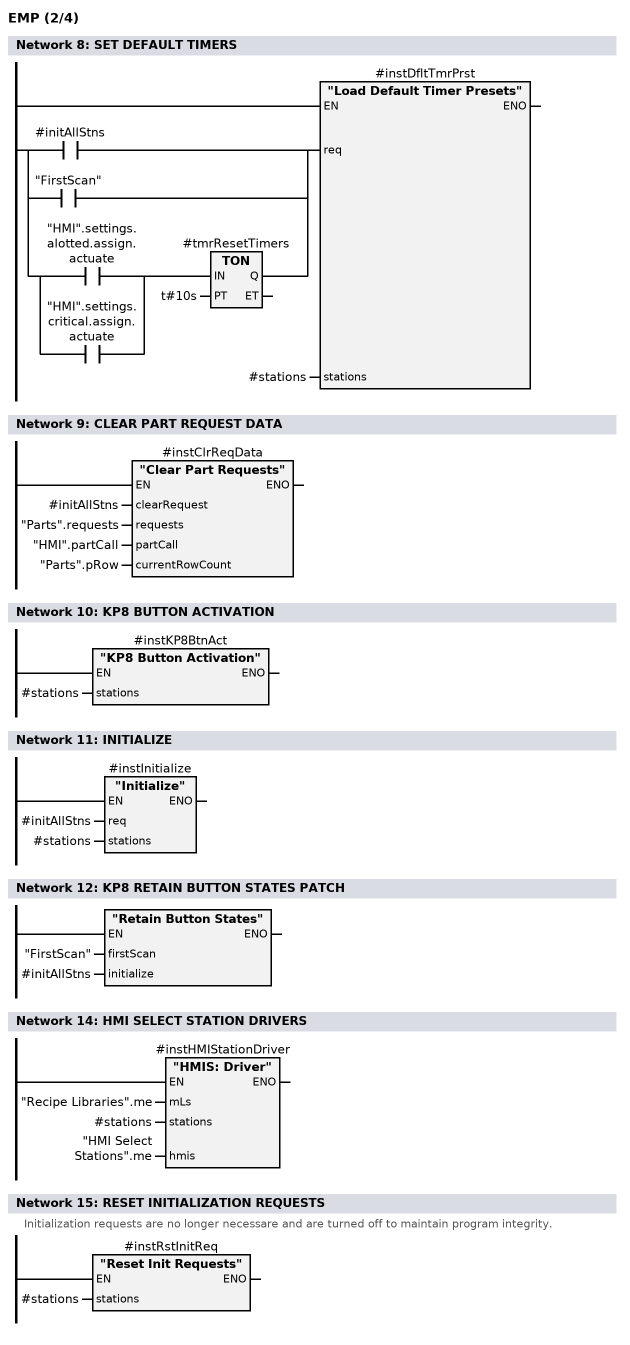
   #tmrResetTimers(IN := "HMI".settings.alotted.assign.actuate OR "HMI".settings.critical.assign.actuate,   // TON
                   PT := t#10s);
   #instDfltTmrPrst(req := #initAllStns OR "FirstScan" OR #tmrResetTimers.Q, stations := #stations);   // "Load Default Timer Presets"
END_REGION

REGION Network 9: CLEAR PART REQUEST DATA
   RUNG wire#powerrail
      #instClrReqData(clearRequest := #initAllStns, requests := "Parts".requests, partCall := "HMI".partCall, currentRowCount := "Parts".pRow)
   END_RUNG
   // the same network as SCL:
   #instClrReqData(clearRequest := #initAllStns,   // "Clear Part Requests"
                   requests := "Parts".requests,
                   partCall := "HMI".partCall,
                   currentRowCount := "Parts".pRow);
END_REGION

REGION Network 10: KP8 BUTTON ACTIVATION
   RUNG wire#powerrail
      #instKP8BtnAct(stations := #stations)
   END_RUNG
   // the same network as SCL:
   #instKP8BtnAct(stations := #stations);   // "KP8 Button Activation"
END_REGION

REGION Network 11: INITIALIZE
   RUNG wire#powerrail
      #instInitialize(req := #initAllStns, stations := #stations)
   END_RUNG
   // the same network as SCL:
   #instInitialize(req := #initAllStns, stations := #stations);   // "Initialize"
END_REGION

REGION Network 12: KP8 RETAIN BUTTON STATES PATCH
   RUNG wire#powerrail
      "Retain Button States"(firstScan := "FirstScan", initialize := #initAllStns)
   END_RUNG
   // the same network as SCL:
   "Retain Button States"(firstScan := "FirstScan", initialize := #initAllStns);
END_REGION

REGION Network 13 (SCL): KP8 DRIVER CALLS
   REGION "LOOP THROUGH STATIONS"
       FOR #i := 0 TO "stnCount" DO
           CASE #i OF
               0..24, 30:
                   #instKP8Drvs[#i](btnIn := #stations.me[#i].kp8In,
                                    hardInit := #stations.me[#i].init.hard,
                                    softInit := #stations.me[#i].init.soft,
                                    btn0Activate := #stations.me[#i].kp8Config.activate[0],
                                    btn0Mode := #stations.me[#i].kp8Config.mode[0],
                                    btn0Group := #stations.me[#i].kp8Config.group[0],
                                    btn0Flash := #stations.me[#i].kp8Config.flash[0],
                                    btn0ColorOn1 := #stations.me[#i].kp8Config.colorOn1[0],
                                    btn0ColorOn2 := #stations.me[#i].kp8Config.colorOn2[0],
                                    btn0ColorOff := #stations.me[#i].kp8Config.colorOff[0],
                                    btn1Activate := #stations.me[#i].kp8Config.activate[1],
                                    btn1Mode := #stations.me[#i].kp8Config.mode[1],
                                    btn1Group := #stations.me[#i].kp8Config.group[1],
                                    btn1Flash := #stations.me[#i].kp8Config.flash[1],
                                    btn1ColorOn1 := #stations.me[#i].kp8Config.colorOn1[1],
                                    btn1ColorOn2 := #stations.me[#i].kp8Config.colorOn2[1],
                                    btn1ColorOff := #stations.me[#i].kp8Config.colorOff[1],
                                    btn2Activate := #stations.me[#i].kp8Config.activate[2],
                                    btn2Mode := #stations.me[#i].kp8Config.mode[2],
                                    btn2Group := #stations.me[#i].kp8Config.group[2],
                                    btn2Flash := #stations.me[#i].kp8Config.flash[2],
                                    btn2ColorOn1 := #stations.me[#i].kp8Config.colorOn1[2],
                                    btn2ColorOn2 := #stations.me[#i].kp8Config.colorOn2[2],
                                    btn2ColorOff := #stations.me[#i].kp8Config.colorOff[2],
                                    btn3Activate := #stations.me[#i].kp8Config.activate[3],
                                    btn3Mode := #stations.me[#i].kp8Config.mode[3],
                                    btn3Group := #stations.me[#i].kp8Config.group[3],
                                    btn3Flash := #stations.me[#i].kp8Config.flash[3],
                                    btn3ColorOn1 := #stations.me[#i].kp8Config.colorOn1[3],
                                    btn3ColorOn2 := #stations.me[#i].kp8Config.colorOn2[3],
                                    btn3ColorOff := #stations.me[#i].kp8Config.colorOff[3],
                                    btn4Activate := #stations.me[#i].kp8Config.activate[4],
                                    btn4Mode := #stations.me[#i].kp8Config.mode[4],
                                    btn4Group := #stations.me[#i].kp8Config.group[4],
                                    btn4Flash := #stations.me[#i].kp8Config.flash[4],
                                    btn4ColorOn1 := #stations.me[#i].kp8Config.colorOn1[4],
                                    btn4ColorOn2 := #stations.me[#i].kp8Config.colorOn2[4],
                                    btn4ColorOff := #stations.me[#i].kp8Config.colorOff[4],
                                    btn5Activate := #stations.me[#i].kp8Config.activate[5],
                                    btn5Mode := #stations.me[#i].kp8Config.mode[5],
                                    btn5Group := #stations.me[#i].kp8Config.group[5],
                                    btn5Flash := #stations.me[#i].kp8Config.flash[5],
                                    btn5ColorOn1 := #stations.me[#i].kp8Config.colorOn1[5],
                                    btn5ColorOn2 := #stations.me[#i].kp8Config.colorOn2[5],
                                    btn5ColorOff := #stations.me[#i].kp8Config.colorOff[5],
                                    btn6Activate := #stations.me[#i].kp8Config.activate[6],
                                    btn6Mode := #stations.me[#i].kp8Config.mode[6],
                                    btn6Group := #stations.me[#i].kp8Config.group[6],
                                    btn6Flash := #stations.me[#i].kp8Config.flash[6],
                                    btn6ColorOn1 := #stations.me[#i].kp8Config.colorOn1[6],
                                    btn6ColorOn2 := #stations.me[#i].kp8Config.colorOn2[6],
                                    btn6ColorOff := #stations.me[#i].kp8Config.colorOff[6],
                                    btn7Activate := #stations.me[#i].kp8Config.activate[7],
                                    btn7Mode := #stations.me[#i].kp8Config.mode[7],
                                    btn7Group := #stations.me[#i].kp8Config.group[7],
                                    btn7Flash := #stations.me[#i].kp8Config.flash[7],
                                    btn7ColorOn1 := #stations.me[#i].kp8Config.colorOn1[7],
                                    btn7ColorOn2 := #stations.me[#i].kp8Config.colorOn2[7],
                                    btn7ColorOff := #stations.me[#i].kp8Config.colorOff[7],
                                    btnStatesOut => #stations.me[#i].btnStates,
                                    btnColorsOut => #stations.me[#i].kp8Out);
               ELSE 
                   ;
           END_CASE;

       END_FOR;
   END_REGION
END_REGION

REGION Network 14: HMI SELECT STATION DRIVERS
   RUNG wire#powerrail
      #instHMIStationDriver(mLs := "Recipe Libraries".me, stations := #stations, hmis := "HMI Select Stations".me)
   END_RUNG
   // the same network as SCL:
   #instHMIStationDriver(mLs := "Recipe Libraries".me, stations := #stations, hmis := "HMI Select Stations".me);   // "HMIS: Driver"
END_REGION

REGION Network 15: RESET INITIALIZATION REQUESTS
   // Initialization requests are no longer necessare and are turned off to maintain program integrity.
   RUNG wire#powerrail
      #instRstInitReq(stations := #stations)
   END_RUNG
   // the same network as SCL:
   #instRstInitReq(stations := #stations);   // "Reset Init Requests"
END_REGION

REGION Network 16: BARCODE SCREEN
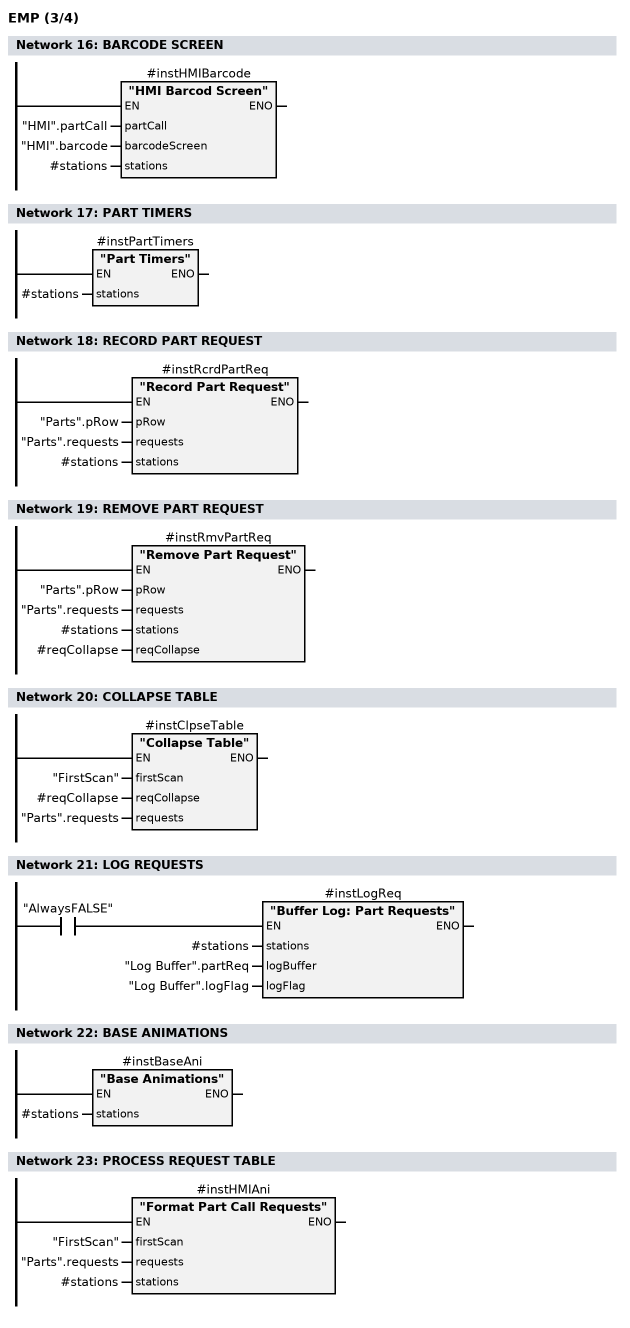
   RUNG wire#powerrail
      #instHMIBarcode(partCall := "HMI".partCall, barcodeScreen := "HMI".barcode, stations := #stations)
   END_RUNG
   // the same network as SCL:
   #instHMIBarcode(partCall := "HMI".partCall, barcodeScreen := "HMI".barcode, stations := #stations);   // "HMI Barcod Screen"
END_REGION

REGION Network 17: PART TIMERS
   RUNG wire#powerrail
      #instPartTimers(stations := #stations)
   END_RUNG
   // the same network as SCL:
   #instPartTimers(stations := #stations);   // "Part Timers"
END_REGION

REGION Network 18: RECORD PART REQUEST
   RUNG wire#powerrail
      #instRcrdPartReq(pRow := "Parts".pRow, requests := "Parts".requests, stations := #stations)
   END_RUNG
   // the same network as SCL:
   #instRcrdPartReq(pRow := "Parts".pRow, requests := "Parts".requests, stations := #stations);   // "Record Part Request"
END_REGION

REGION Network 19: REMOVE PART REQUEST
   RUNG wire#powerrail
      #instRmvPartReq(pRow := "Parts".pRow, requests := "Parts".requests, stations := #stations, reqCollapse := #reqCollapse)
   END_RUNG
   // the same network as SCL:
   #instRmvPartReq(pRow := "Parts".pRow,   // "Remove Part Request"
                   requests := "Parts".requests,
                   stations := #stations,
                   reqCollapse := #reqCollapse);
END_REGION

REGION Network 20: COLLAPSE TABLE
   RUNG wire#powerrail
      #instClpseTable(firstScan := "FirstScan", reqCollapse := #reqCollapse, requests := "Parts".requests)
   END_RUNG
   // the same network as SCL:
   #instClpseTable(firstScan := "FirstScan", reqCollapse := #reqCollapse, requests := "Parts".requests);   // "Collapse Table"
END_REGION

REGION Network 21: LOG REQUESTS
   RUNG wire#powerrail
      Contact( "AlwaysFALSE" )
      #instLogReq(stations := #stations, logBuffer := "Log Buffer".partReq, logFlag := "Log Buffer".logFlag)
   END_RUNG
   // the same network as SCL:
   IF "AlwaysFALSE" THEN
       #instLogReq(stations := #stations, logBuffer := "Log Buffer".partReq, logFlag := "Log Buffer".logFlag);   // "Buffer Log: Part Requests"
   END_IF;
END_REGION

REGION Network 22: BASE ANIMATIONS
   RUNG wire#powerrail
      #instBaseAni(stations := #stations)
   END_RUNG
   // the same network as SCL:
   #instBaseAni(stations := #stations);   // "Base Animations"
END_REGION

REGION Network 23: PROCESS REQUEST TABLE
   RUNG wire#powerrail
      #instHMIAni(firstScan := "FirstScan", requests := "Parts".requests, stations := #stations)
   END_RUNG
   // the same network as SCL:
   #instHMIAni(firstScan := "FirstScan", requests := "Parts".requests, stations := #stations);   // "Format Part Call Requests"
END_REGION

REGION Network 24: HMI POPULATE TABLE
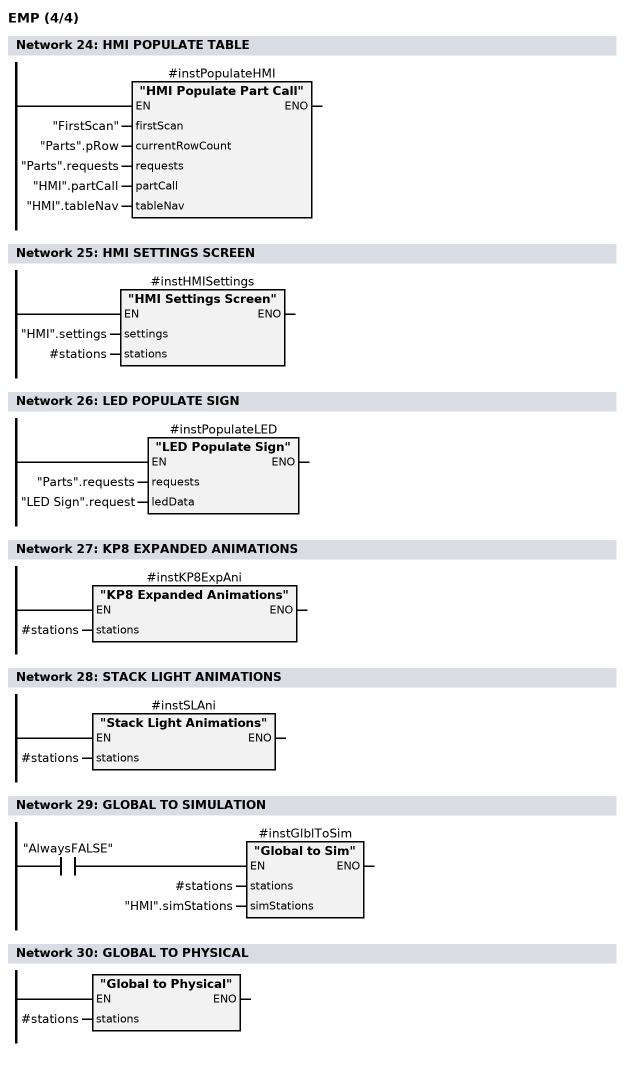
   RUNG wire#powerrail
      #instPopulateHMI(firstScan := "FirstScan", currentRowCount := "Parts".pRow, requests := "Parts".requests, partCall := "HMI".partCall, tableNav := "HMI".tableNav)
   END_RUNG
   // the same network as SCL:
   #instPopulateHMI(firstScan := "FirstScan",   // "HMI Populate Part Call"
                    currentRowCount := "Parts".pRow,
                    requests := "Parts".requests,
                    partCall := "HMI".partCall,
                    tableNav := "HMI".tableNav);
END_REGION

REGION Network 25: HMI SETTINGS SCREEN
   RUNG wire#powerrail
      #instHMISettings(settings := "HMI".settings, stations := #stations)
   END_RUNG
   // the same network as SCL:
   #instHMISettings(settings := "HMI".settings, stations := #stations);   // "HMI Settings Screen"
END_REGION

REGION Network 26: LED POPULATE SIGN
   RUNG wire#powerrail
      #instPopulateLED(requests := "Parts".requests, ledData := "LED Sign".request)
   END_RUNG
   // the same network as SCL:
   #instPopulateLED(requests := "Parts".requests, ledData := "LED Sign".request);   // "LED Populate Sign"
END_REGION

REGION Network 27: KP8 EXPANDED ANIMATIONS
   RUNG wire#powerrail
      #instKP8ExpAni(stations := #stations)
   END_RUNG
   // the same network as SCL:
   #instKP8ExpAni(stations := #stations);   // "KP8 Expanded Animations"
END_REGION

REGION Network 28: STACK LIGHT ANIMATIONS
   RUNG wire#powerrail
      #instSLAni(stations := #stations)
   END_RUNG
   // the same network as SCL:
   #instSLAni(stations := #stations);   // "Stack Light Animations"
END_REGION

REGION Network 29: GLOBAL TO SIMULATION
   RUNG wire#powerrail
      Contact( "AlwaysFALSE" )
      #instGlblToSim(stations := #stations, simStations := "HMI".simStations)
   END_RUNG
   // the same network as SCL:
   IF "AlwaysFALSE" THEN
       #instGlblToSim(stations := #stations, simStations := "HMI".simStations);   // "Global to Sim"
   END_IF;
END_REGION

REGION Network 30: GLOBAL TO PHYSICAL
   RUNG wire#powerrail
      "Global to Physical"(stations := #stations)
   END_RUNG
   // the same network as SCL:
   "Global to Physical"(stations := #stations);
END_REGION
END_FUNCTION_BLOCK

FUNCTION "Retain Button States" : Void   // FC36, SCL
{ S7_Optimized_Access := 'TRUE' }
VERSION : 0.1
   VAR_INPUT
      firstScan : Bool;
      initialize : Bool;
   END_VAR
   VAR_TEMP
      i : Int;
      j : Int;
   END_VAR
BEGIN
   FOR #i := 0 TO "stnCount" DO
           FOR #j := 0 TO "ptsPerStn" DO
               IF #firstScan THEN
                   "EMP IDB".instKP8Drvs[#i].btnStateArrayInt[#j] :=
                   "EMP IDB".stations.me[#i].btnStates[#j];
               END_IF;
               IF #initialize THEN
                   "EMP IDB".instKP8Drvs[#i].btnStateArrayInt[#j] := FALSE;
                   "EMP IDB".stations.me[#i].btnStates[#j] := FALSE;
               END_IF;
           END_FOR;
   END_FOR;
END_FUNCTION

ORGANIZATION_BLOCK "Main"   // OB1, LAD, ProgramCycle
TITLE = "Main Program Sweep (Cycle)"
{ S7_Optimized_Access := 'TRUE' }
VERSION : 0.1
   VAR_INPUT
      Initial_Call : Bool;   // Initial call of this OB
      Remanence : Bool;   // =True, if remanent data are available
   END_VAR
BEGIN

REGION Network 1
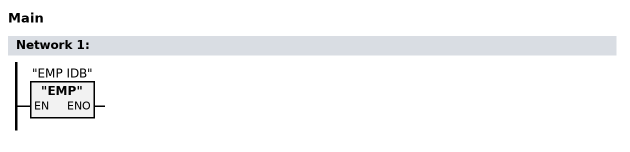
   RUNG wire#powerrail
      "EMP IDB"()
   END_RUNG
   // the same network as SCL:
   "EMP IDB"();   // "EMP"
END_REGION
END_ORGANIZATION_BLOCK

// folder: Global/Physical

FUNCTION "Physical to Global" : Void   // FC1, LAD
{ S7_Optimized_Access := 'TRUE' }
VERSION : 0.1
   VAR_IN_OUT
      stations : "Stations";
   END_VAR
   VAR_TEMP
      i : Int;
      kp8In : DWord;
   END_VAR
BEGIN

REGION Network 1 (SCL): MAIN LOOP
   FOR #i := 0 TO "stnCount" DO

       CASE #i OF
           "VOLVO 16 01":
               #kp8In := "VOLVO 16 01 KP8 In";
           "VOLVO 16 02":
               #kp8In := "VOLVO 16 02 KP8 In";
           "VOLVO 16 03":
               #kp8In := "VOLVO 16 03 KP8 In";
           "VOLVO 16 04":
               #kp8In := "VOLVO 16 04 KP8 In";
           "VOLVO 16 05":
               #kp8In := "VOLVO 16 05 KP8 In";
           "VOLVO 16 06":
               #kp8In := "VOLVO 16 06 KP8 In";
           "VOLVO 16 07":
               #kp8In := "VOLVO 16 07 KP8 In";
           "VOLVO 16 08":
               #kp8In := "VOLVO 16 08 KP8 In";
           "VOLVO 16 09":
               #kp8In := "VOLVO 16 09 KP8 In";
           "VOLVO 16 10":
               #kp8In := "VOLVO 16 10 KP8 In";
           "VOLVO 16 11":
               #kp8In := "VOLVO 16 11 KP8 In";
           "CHM 01":
               #kp8In := "CHM 01 KP8 In";
           "CHM 02":
               #kp8In := "CHM 02 KP8 In";
           "CHM 03":
               #kp8In := "CHM 03 KP8 In";
           "CHM 04":
               #kp8In := "CHM 04 KP8 In";
           "CHM 05":
               #kp8In := "CHM 05 KP8 In";
           "CDO 01":
               #kp8In := "CDO 01 KP8 In";
           "CDO 02":
               #kp8In := "CDO 02 KP8 In";
           "CDO 03":
               #kp8In := "CDO 03 KP8 In";
           "BFL 01":
               #kp8In := "BFL 01 KP8 In";
           "BFL 02":
               #kp8In := "BFL 02 KP8 In";
           "BFL 03":
               #kp8In := "BFL 03 KP8 In";
           "LGS 01":
               #kp8In := "LGS 01 KP8 In";
           "LGS 02":
               #kp8In := "LGS 02 KP8 In";
           "LGS 03":
               #kp8In := "LGS 03 KP8 In";
           "CV 01":
               #kp8In := "CV 01 KP8 In";
           "CV 02":
               #kp8In := "CV 02 KP8 In";
           "CV 03":
               #kp8In := "CV 03 KP8 In";
           "CV 04":
               #kp8In := "CV 04 KP8 In";
           "PC 01":
               #kp8In := "PC 01 KP8 In"; 
           "PC 02":
               #kp8In := "PC 02 KP8 In";
       END_CASE;

       #stations.me[#i].kp8In := #kp8In.%B3;

   END_FOR;
END_REGION
END_FUNCTION

FUNCTION "Global to Physical" : Void   // FC5, LAD
{ S7_Optimized_Access := 'TRUE' }
VERSION : 0.1
   VAR_IN_OUT
      stations : "Stations";
   END_VAR
   VAR_TEMP
      i : Int;
      j : Int;
      IO : DWord;
      "KP8 In" : DWord;
      "KP8 Out" : DWord;
      Card : Int;
      stnCount : Int;
   END_VAR
BEGIN

REGION Network 1 (SCL): MAIN LOOP
   FOR #i := 0 TO "stnCount" DO

       #IO := #stations.me[#i].stackLightOut;
       #"KP8 Out" := #stations.me[#i].kp8Out;

       CASE #i OF
           "VOLVO 16 01":
               "VOLVO 16 01 IO" := #IO;
               "VOLVO 16 01 KP8 Out" := #"KP8 Out";
           "VOLVO 16 02":
               "VOLVO 16 02 IO" := #IO;
               "VOLVO 16 02 KP8 Out" := #"KP8 Out";
           "VOLVO 16 03":
               "VOLVO 16 03 IO" := #IO;
               "VOLVO 16 03 KP8 Out" := #"KP8 Out";
           "VOLVO 16 04":
               "VOLVO 16 04 IO" := #IO;
               "VOLVO 16 04 KP8 Out" := #"KP8 Out";
           "VOLVO 16 05":
               "VOLVO 16 05 IO" := #IO;
               "VOLVO 16 05 KP8 Out" := #"KP8 Out";
           "VOLVO 16 06":
               "VOLVO 16 06 IO" := #IO;
               "VOLVO 16 06 KP8 Out" := #"KP8 Out";
           "VOLVO 16 07":
               "VOLVO 16 07 IO" := #IO;
               "VOLVO 16 07 KP8 Out" := #"KP8 Out";
           "VOLVO 16 08":
               "VOLVO 16 08 IO" := #IO;
               "VOLVO 16 08 KP8 Out" := #"KP8 Out";
           "VOLVO 16 09":
               "VOLVO 16 09 IO" := #IO;
               "VOLVO 16 09 KP8 Out" := #"KP8 Out";
           "VOLVO 16 10":
               "VOLVO 16 10 IO" := #IO;
               "VOLVO 16 10 KP8 Out" := #"KP8 Out";
           "VOLVO 16 11":
               "VOLVO 16 11 IO" := #IO;
               "VOLVO 16 11 KP8 Out" := #"KP8 Out";
           "CHM 01":
               "CHM 01 IO" := #IO;
               "CHM 01 KP8 Out" := #"KP8 Out";
           "CHM 02":
               "CHM 02 IO" := #IO;
               "CHM 02 KP8 Out" := #"KP8 Out";
           "CHM 03":
               "CHM 03 IO" := #IO;
               "CHM 03 KP8 Out" := #"KP8 Out";
           "CHM 04":
               "CHM 04 IO" := #IO;
               "CHM 04 KP8 Out" := #"KP8 Out";
           "CHM 05":
               "CHM 05 IO" := #IO;
               "CHM 05 KP8 Out" := #"KP8 Out";
           "CDO 01":
               "CDO 01 IO" := #IO;
               "CDO 01 KP8 Out" := #"KP8 Out";
           "CDO 02":
               "CDO 02 IO" := #IO;
               "CDO 02 KP8 Out" := #"KP8 Out";
           "CDO 03":
               "CDO 03 IO" := #IO;
               "CDO 03 KP8 Out" := #"KP8 Out";
           "BFL 01":
               "BFL 01 IO" := #IO;
               "BFL 01 KP8 Out" := #"KP8 Out";
           "BFL 02":
               "BFL 02 IO" := #IO;
               "BFL 02 KP8 Out" := #"KP8 Out";
           "BFL 03":
               "BFL 03 IO" := #IO;
               "BFL 03 KP8 Out" := #"KP8 Out";
           "LGS 01":
               "LGS 01 IO" := #IO;
               "LGS 01 KP8 Out" := #"KP8 Out";
           "LGS 02":
               "LGS 02 IO" := #IO;
               "LGS 02 KP8 Out" := #"KP8 Out";
           "LGS 03":
               "LGS 03 IO" := #IO;
               "LGS 03 KP8 Out" := #"KP8 Out";
           "CV 01":
               "CV 01 IO" := #IO;
               "CV 01 KP8 Out" := #"KP8 Out";
           "CV 02":
               "CV 02 IO" := #IO;
               "CV 02 KP8 Out" := #"KP8 Out";
           "CV 03":
               "CV 03 IO" := #IO;
               "CV 03 KP8 Out" := #"KP8 Out";
           "CV 04":
               "CV 04 IO" := #IO;
               "CV 04 KP8 Out" := #"KP8 Out";
           "PC 01":
               "PC 01 IO" := #IO;
               "PC 01 KP8 Out" := #"KP8 Out";
           "PC 02":
               "PC 02 IO" := #IO;
               "PC 02 KP8 Out" := #"KP8 Out";

       END_CASE;

   END_FOR;
END_REGION
END_FUNCTION

// folder: HMI Stations

FUNCTION_BLOCK "HMIS: Driver"   // FB32, LAD
{ S7_Optimized_Access := 'TRUE' }
VERSION : 0.1
   VAR_INPUT
      mLs : "Recipe: Libraries";
   END_VAR
   VAR_IN_OUT
      stations : "Stations";
      hmis : Array[0.."hmiStnCount"] of "HSS: Compressed";
   END_VAR
   VAR
      recipeSelector : Array[0.."hmiStnCount"] of Int;
      r1 : Array[0.."hmiStnCount"] of DInt;
      instsHSSMenuSelect : Array[0.."hmiStnCount"] of "HMIS: Recipe Selection";
      instsHSSPartSelect : Array[0.."hmiStnCount"] of "HMIS: Part Selection";
   END_VAR
   VAR_TEMP
      i : Int;
   END_VAR
   VAR CONSTANT
      hssOffset : Int := 25;
   END_VAR
BEGIN

REGION Network 1 (SCL): TEMPLATE SCREENS
   FOR #i := 0 TO "hmiStnCount" DO
       "HMIS: Template"(menuLibrary := #mLs.stations[#i + #hssOffset],
                       menuSelector := #recipeSelector[#i],
                       tmplt := #hmis[#i].scrnTmplt);
       #instsHSSMenuSelect[#i](lib := #mLs.stations[#i + #hssOffset],
                               slctScreen := #hmis[#i].scrnSlctMn,
                               r1 := #r1[#i],
                               station := #stations.me[#i + #hssOffset],
                               recipeSelector := #recipeSelector[#i]);
       #instsHSSPartSelect[#i](recipeNum:= #recipeSelector[#i],
                              lib:=#mLs.stations[#i + #hssOffset],
                              slctScreen:=#hmis[#i].scrnSlctPrt,
                              station:=#stations.me[#i + #hssOffset]);

   END_FOR;
END_REGION
END_FUNCTION_BLOCK

FUNCTION_BLOCK "HMIS: Part Selection"   // FB33, SCL
{ S7_Optimized_Access := 'TRUE' }
VERSION : 0.1
   VAR_INPUT
      recipeNum : Int;
      lib : "Recipe: Library";
   END_VAR
   VAR_IN_OUT
      slctScreen : "HSS: Part Selection Screen";
      station : "Station";
   END_VAR
   VAR
      oldBtnsIn : Array[0..31] of Bool;
   END_VAR
   VAR_TEMP
      eval : "HSS: Part Selection Screen";
      i : Int;
      btnsIn : Array[0..31] of Bool;
      btnStates : Array[0.."ptsPerStn"] of Bool;
   END_VAR
BEGIN
   #eval := #slctScreen;


   SCATTER(IN := #slctScreen.pbs ,
           OUT => #btnsIn);
   #btnStates := #station.btnStates;


   FOR #i := 0 TO "ptsPerStn" DO
       IF #btnsIn[#i] AND #btnsIn[#i] <> #oldBtnsIn[#i] THEN
           #btnStates[#i] := NOT #btnStates[#i];
       END_IF;
   END_FOR;


   FOR #i := 0 TO "ptsPerStn" DO
       "Part Select Button"(recipeNum := #recipeNum,
                            lib := #lib,
                            actuate := #btnsIn[#i],
                            btnNum := #i,
                            stn:= #station,
                            partSelectScreen := #eval);
   END_FOR;


   #station.btnStates := #btnStates;
   #oldBtnsIn := #btnsIn;
   #slctScreen := #eval;
END_FUNCTION_BLOCK

FUNCTION_BLOCK "HMIS: Recipe Selection"   // FB35, SCL
{ S7_Optimized_Access := 'TRUE' }
VERSION : 0.1
   VAR_INPUT
      lib : "Recipe: Library";
   END_VAR
   VAR_IN_OUT
      slctScreen : "HSS: Menu Selection Screen";
      r1 : DInt;
      recipeSelector : Int;
      station : "Station";
   END_VAR
   VAR
      old : Struct
         navPress : Bool;
      END_STRUCT;
      instTableNavigation : "Table Navigatio";
   END_VAR
   VAR_TEMP
      eval : "HSS: Menu Selection Screen";
      pbs : Array[0..#pbFlagCnt] of Bool;
      POS : DInt;
      status : DInt;
      i : Int;
      btnNum : Int;
      pRowVisLbl : Int;
      pRowInvisLbl : Int;
      pRecipeInvisLbl : Int;
      pRecipeVisLbl : Int;
      pRecipeLib : Int;
      pRowTxt : Int;
      pRecipeTxt : Int;
      shifter : DWord;
      btnsAsBool : Array[0..31] of Bool;
      rows : Array[0..99] of DInt;
      offset : DInt;
      navPress : Bool;
      selPress : Bool;
      maxRows : DInt;
      tmrReal : Real;
      partNumber : WString;
   END_VAR
   VAR CONSTANT
      pbFlagCnt : Int := 31;
      btnCnt : Int := 5;
      navMask : DWord := 16#0000_003F;
      visRows : DInt := 6;
      home : DInt := -1000;
      end : DInt := -2000;
      alotted : Real := 1800.0;
      critical : Real := 300.0;
   END_VAR
BEGIN
   REGION "INITITALIZE LOCALS"

       #eval := #slctScreen;
       #maxRows := #lib.size;
       SCATTER(IN := #eval.pbs,
               OUT => #btnsAsBool);

   END_REGION


   REGION "GET RECIPE SELECTION PRESS" 

       REGION "GET RECIPE SELECTOR NUMBER"

           FOR #i := 6 TO 31 DO
               IF #btnsAsBool[#i] THEN

                   #recipeSelector := DINT_TO_INT(#r1) + #i - 6;

                   IF #recipeSelector > #maxRows -1 THEN
                       #recipeSelector := #recipeSelector - DINT_TO_INT(#maxRows);
                   END_IF;

                   IF #recipeSelector < 0 THEN
                       #recipeSelector := DINT_TO_INT(#maxRows) + #recipeSelector;
                   END_IF;

                   #selPress := TRUE;
                   EXIT;
               END_IF;
           END_FOR;

       END_REGION


       FOR #i := 0 TO "ptsPerStn" DO
           #station.partNumbers[#i] := #lib.raw[#recipeSelector, #i];
           IF #i = 1 THEN
               #station.partNumbers[#i] := WSTRING#'DUNNAGE';
           END_IF;

       END_FOR;

       REGION "SET DEFAULT TIMERS"
           FOR #i := 0 TO "ptsPerStn" DO

               REGION "COPY TO LOCAL"
                   #partNumber := #station.partNumbers[#i];
               END_REGION

               REGION "IF BUTTON HAS ASSOCIATED PN"
                   IF LEN(#partNumber) <> 0 THEN

                       REGION "COPY TO LOCAL"
                           #tmrReal := #station.presetTime.allotted[#i];
                       END_REGION

                       REGION "ON NO TIME ENTERED"
                           IF #tmrReal = 0.0 THEN

                               REGION "ASSIGN ALLOTTED VALUES"
                                   #station.presetTime.allotted[#i] := #alotted;
                               END_REGION

                           END_IF;
                       END_REGION

                       REGION "COPY TO LOCAL"
                           #tmrReal := #station.presetTime.critical[#i];
                       END_REGION

                       REGION "ON NO TIME ENTERED"
                           IF #tmrReal = 0.0 THEN

                               REGION "ASSIGN CRITICAL VALUES"
                                   #station.presetTime.critical[#i] := #critical;
                               END_REGION

                           END_IF;
                       END_REGION

                   END_IF;
               END_REGION

               REGION "IF BUTTON HAS NO ASSOCIATED PN"
                   IF LEN(#partNumber) = 0 THEN

                       REGION "COPY TO LOCAL"
                           #tmrReal := #station.presetTime.allotted[#i];
                       END_REGION

                       REGION "ON NO TIME ENTERED"
                           IF #tmrReal <> 0.0 THEN

                               REGION "ASSIGN ALLOTTED VALUES"
                                   #station.presetTime.allotted[#i] := 0.0;
                               END_REGION

                           END_IF;
                       END_REGION

                       REGION "COPY TO LOCAL"
                           #tmrReal := #station.presetTime.critical[#i];
                       END_REGION

                       REGION "ON NO TIME ENTERED"
                           IF #tmrReal <> 0.0 THEN

                               REGION "ASSIGN CRITICAL VALUES"
                                   #station.presetTime.critical[#i] := 0.0;
                               END_REGION

                           END_IF;
                       END_REGION

                   END_IF;
               END_REGION


           END_FOR;
       END_REGION

   END_REGION


   REGION "TABLE NAVIGATION"
       IF #maxRows > #visRows THEN
           IF #eval.pbs.%X0 THEN
               #offset := #home;
           END_IF;
           IF #eval.pbs.%X1 THEN
               #offset := -1 * #visRows;
           END_IF;
           IF #eval.pbs.%X2 THEN
               #offset := -1;
           END_IF;
           IF #eval.pbs.%X3 THEN
               #offset := 1;
           END_IF;
           IF #eval.pbs.%X4 THEN
               #offset := #visRows;
           END_IF;
           IF #eval.pbs.%X5 THEN
               #offset := #end;
           END_IF;

           IF (#eval.pbs AND #navMask) <> 0 THEN
               #navPress := true;
           END_IF;

           #instTableNavigation(maxRows := #maxRows,
                                visRows := #visRows,
                                offset := #offset,
                                trigger := #navPress,
                                r1 := #r1,
                                rowIndices := #rows);
       END_IF;

       IF #maxRows <= #visRows THEN
           FOR #i := 0 TO #visRows - 1 DO
               #rows[#i] := #i;
           END_FOR;
       END_IF;

   END_REGION


   REGION "NAV BUTTONS"

       FOR #i := 0 TO #visRows - 1 DO
           "Recipe Nav Button"(visRows := DINT_TO_INT(#visRows),
                               actuate := #btnsAsBool[#i],
                               maxRows := DINT_TO_INT(#maxRows),
                               btnNum := #i,
                               recipeSelectScreen := #eval);
       END_FOR;

   END_REGION



   REGION "RECIPE SELECT BUTTONS"

       IF (#navPress AND NOT #old.navPress) OR
           (#maxRows <= #visRows) THEN

           FOR #i := 0 TO #visRows - 1 DO
               "Recipe Select Button"(visRows := DINT_TO_INT(#visRows),
                                      rowNum := DINT_TO_INT(#rows[#i]),
                                      lib := #lib,
                                      actuate := #btnsAsBool[#i + 6],
                                      maxRows := DINT_TO_INT(#maxRows),
                                      btnNum := #i,
                                      recipeSelectScreen := #eval);
           END_FOR;
       END_IF;

   END_REGION


   REGION "CHANGE DETECTION"

       #old.navPress := #navPress;

   END_REGION


   REGION "COPY TO GLOBAL"

       #slctScreen := #eval;

   END_REGION
END_FUNCTION_BLOCK

FUNCTION "HMIS: Template" : Void   // FC24, SCL
{ S7_Optimized_Access := 'TRUE' }
VERSION : 0.1
   VAR_INPUT
      menuLibrary : "Recipe: Library";
      menuSelector : Int;
   END_VAR
   VAR_IN_OUT
      tmplt : "HSS: Template Screen";
   END_VAR
   VAR_TEMP
      i : Int;
   END_VAR
BEGIN
   #tmplt.animate[0] := "BgGray";
   #tmplt.text[0] := "Word Wrap"(stringIn := #menuLibrary.wip[#menuSelector],
                                 maxLength := 22);
END_FUNCTION

FUNCTION "Recipe Select Button" : Void   // FC31, SCL
{ S7_Optimized_Access := 'TRUE' }
VERSION : 0.1
   VAR_INPUT
      visRows : Int;
      rowNum : Int;
      lib : "Recipe: Library";
      actuate : Bool;
      maxRows : Int;
      btnNum : Int;
   END_VAR
   VAR_IN_OUT
      recipeSelectScreen : "HSS: Menu Selection Screen";
   END_VAR
   VAR_TEMP
      eval : "HSS: Menu Selection Screen";
      pRowVisLbl : Int;
      pRowInvisLbl : Int;
      pRowTxt : Int;
      pRecipeTxt : Int;
      maxLen : Int;
   END_VAR
BEGIN
   REGION "COPY TO LOCAL"
       #eval := #recipeSelectScreen;
   END_REGION


   REGION "NARROW"
       IF #maxRows > #visRows THEN
           #pRowVisLbl := #btnNum + #visRows;
           #pRowInvisLbl := #btnNum + (3 * #visRows);
           #maxLen := 22;
       END_IF;
   END_REGION


   REGION "WIDE"
       IF #maxRows <= #visRows THEN
           #pRowVisLbl := #btnNum + (3 * #visRows);
           #pRowInvisLbl := #btnNum + #visRows + 1;
           #maxLen := 28;
       END_IF;
   END_REGION


   REGION "ROW COUNT INDEPENDENT"
       #pRowTxt := (#btnNum * 2) + #visRows;
       #pRecipeTxt := #pRowTxt + 1;
   END_REGION


   REGION "DRAW"
       IF #btnNum < #maxRows THEN
           #eval.animate[#pRowVisLbl] := "BgGray";
       END_IF;
       IF #btnNum >= #maxRows THEN
           #eval.animate[#pRowVisLbl] := "invisible";
       END_IF;
       #eval.animate[#pRowInvisLbl] := "invisible";
       #eval.txt[#pRowTxt] := "Strip Sign"(DINT_TO_WSTRING(#rowNum));
       #eval.txt[#pRecipeTxt] := "Word Wrap"(stringIn := #lib.wip[#rowNum],
                                             maxLength := #maxLen);
   END_REGION

   REGION "ACTUATION ANIMATION"
       IF #actuate THEN
           #eval.animate[#pRowVisLbl] := "BgLTe";
       END_IF;
   END_REGION


   REGION "COPY TO GLOBAL"
       #recipeSelectScreen := #eval;
   END_REGION
END_FUNCTION

FUNCTION "Part Select Button" : Void   // FC34, SCL
{ S7_Optimized_Access := 'TRUE' }
VERSION : 0.1
   VAR_INPUT
      recipeNum : Int;
      lib : "Recipe: Library";
      actuate : Bool;
      btnNum : Int;
      stn : "Station";
   END_VAR
   VAR_IN_OUT
      partSelectScreen : "HSS: Part Selection Screen";
   END_VAR
   VAR_TEMP
      eval : "HSS: Part Selection Screen";
      i : Int;
      target : Int;
   END_VAR
   VAR CONSTANT
      blank : WString;
      anDefault : USInt := 0;
      anRequested : USInt := 1;
      anSolidRed : USInt := 2;
      anFlashRed : USInt := 3;
      anPartOrdered : USInt := 4;
   END_VAR
BEGIN
   REGION "COPY TO LOCAL"
       #eval := #partSelectScreen;
   END_REGION


   REGION "DRAW NEEDED BUTTONS"
       IF #stn.partNumbers[#btnNum] = #blank THEN
           #eval.animate[#btnNum] := "invisible";
       END_IF;
       IF #stn.partNumbers[#btnNum] <> #blank THEN
           CASE #stn.animations[#btnNum] OF
               #anDefault:
                   #eval.animate[#btnNum] := "BgLGr";
               #anRequested:
                   #eval.animate[#btnNum] := "BgDYe";
               #anSolidRed:
                   #eval.animate[#btnNum] := "BgDRd";
               #anFlashRed:
                   #eval.animate[#btnNum] := "FlDrd";
               #anPartOrdered:
                   #eval.animate[#btnNum] := "BgDBl";
               ELSE:
                   ;
           END_CASE;
       END_IF;
   END_REGION


   REGION "ACTUATION ANIMATION"
       IF #actuate THEN
           #eval.animate[#btnNum] := "BgLTe";
       END_IF;
   END_REGION


   REGION "PART NUMBER"
       #eval.txt[#btnNum] :=#stn.partNumbers[#btnNum];
   END_REGION


   REGION "COPY TO GLOBAL"
       #partSelectScreen := #eval;
   END_REGION
END_FUNCTION

// folder: Other OBs

ORGANIZATION_BLOCK "Rack or station failure"   // OB86, LAD, RackStationFailure
{ S7_Optimized_Access := 'TRUE' }
VERSION : 0.1
   VAR_INPUT
      LADDR : Hw_Device;   // Hardware identifier
      Event_Class : Byte;   // Event class
      Fault_ID : Byte;   // Fault identifier
   END_VAR
BEGIN
END_ORGANIZATION_BLOCK

ORGANIZATION_BLOCK "Programming error"   // OB121, LAD, ProgrammingError
{ S7_Optimized_Access := 'TRUE' }
VERSION : 0.1
   VAR_INPUT
      BlockNr : UInt;   // Number of causing block
      Reaction : USInt;   // 0:ignore, 1:substitute, 2:skip
      Fault_ID : Byte;   // Fault identifier
      BlockType : USInt;   // 16#01:OB, 16#02:FC, 16#03:FB, 16#04:SFC, 16#05:SFB, 16#06:DB: Type of block causing the error
      Area : USInt;   // Area where the error occured
      DBNr : DB_ANY;   // DB number if Area = DB or DI
      Csg_OBNr : OB_Any;   // Number of OB causing the error
      Csg_Prio : USInt;   // Priority of OB causing the error
      Width : USInt;   // 0:bit, 1:byte, 2:word, 3:dword, 4:lword
   END_VAR
BEGIN
END_ORGANIZATION_BLOCK

ORGANIZATION_BLOCK "IO access error"   // OB122, LAD, IOAccessError
{ S7_Optimized_Access := 'TRUE' }
VERSION : 0.1
   VAR_INPUT
      BlockNr : UInt;   // Number of causing block
      Reaction : USInt;   // 0:ignore, 1:substitute, 2:skip
      Fault_ID : Byte;   // 16#42:reading, 16#43:writing
      BlockType : USInt;   // 16#01:OB, 16#02:FC, 16#03:FB, 16#04:SFC, 16#05:SFB, 16#06:DB: Type of block causing the error
      Area : USInt;   // 16#81:I, 16#82:Q: IO area where the IOaccess error occured
      DBNr : DB_ANY;   // Reserved for system
      Csg_OBNr : OB_Any;   // Number of OB causing the error
      Csg_Prio : USInt;   // Priority of OB causing the error
      Width : USInt;   // 0:bit, 1:byte, 2:word, 3:dword, 4:lword
   END_VAR
BEGIN
END_ORGANIZATION_BLOCK

// folder: Part Request

FUNCTION_BLOCK "Record Part Request"   // FB6, SCL
{ S7_Optimized_Access := 'TRUE' }
VERSION : 0.1
   VAR_IN_OUT
      pRow : Int;
      requests : "Part Request Data";
      stations : "Stations";
   END_VAR
   VAR
      enterAddress : Bool;
      old : Struct
         presses : "Station Old Presses";
      END_STRUCT;
   END_VAR
   VAR_TEMP
      address : UInt;
      hasPart : Bool;
      i : Int;
      j : Int;
      k : Int;
      logAddress : UInt;
      noPart : Bool;
      oldPartReq : Bool;
      partReq : Bool;
      partNumber : WString;
   END_VAR
BEGIN
   REGION "FOR EACH STATION"
       FOR #i := 0 TO "stnCount" DO

           REGION "FOR EACH BUTTON"
               // j = 0 is excluded because it is used as a station reset button
               FOR #j := 1 TO "ptsPerStn" DO

                   REGION "COPY TO LOCAL"
                       #partReq := #stations.me[#i].btnStates[#j];
                       #oldPartReq := #old.presses.me[#i,#j];
                   END_REGION

                   REGION "DETERMINE STATE"

                       REGION "ON NEW REQUEST"
                           IF #partReq AND NOT #oldPartReq THEN

                               REGION "COPY TO LOCAL"
                                   #partNumber := #stations.me[#i].partNumbers[#j];
                               END_REGION

                               REGION "BUTTON HAS NO PN"
                                   IF LEN(#partNumber) = 0 THEN
                                       #hasPart := FALSE;
                                       #noPart := TRUE;
                                   END_IF;
                               END_REGION

                               REGION "BUTTON HAS PN"
                                   IF LEN(#partNumber) <> 0 THEN
                                       #hasPart := TRUE;
                                       #noPart := FALSE;
                                   END_IF;
                               END_REGION

                           END_IF;

                           REGION "SAVE FOR CHANGE DETECTION"
                               #old.presses.me[#i, #j] := #stations.me[#i].btnStates[#j];
                           END_REGION

                       END_REGION

                   END_REGION

                   REGION "NO PART"
                       IF #noPart THEN

                           REGION "TURN OFF THE LIGHTS"
                               #hasPart := FALSE;
                               #noPart := FALSE;
                               #enterAddress := FALSE;
                           END_REGION

                       END_IF;
                   END_REGION

                   REGION "HAS PART"
                       IF #hasPart THEN

                           REGION "TURN OFF THE LIGHTS"
                               #hasPart := FALSE;
                               #noPart := FALSE;
                               #enterAddress := FALSE;
                           END_REGION

                           REGION "CALCULATE ADDRESS"
                               #address := (INT_TO_UINT(#i) + 1) * 10 + (INT_TO_UINT(#j) + 1);
                           END_REGION

                           REGION "SET FLAG"
                               #enterAddress := TRUE;
                           END_REGION

                           REGION "CHECK FOR ENTRY IN DB"
                               REGION "FOR EACH ROW IN PART DB"
                                   FOR #k := 0 TO "partReqDataRowCount" DO

                                       REGION "COPY TO LOCAL"
                                           #logAddress := #requests.row[#k].address;
                                       END_REGION

                                       REGION "RESET FLAG"
                                           IF #logAddress = #address THEN
                                               #enterAddress := FALSE;
                                           END_IF;
                                       END_REGION

                                   END_FOR;
                               END_REGION
                           END_REGION


                       END_IF;
                   END_REGION

                   REGION "SAVE ROW DATA"
                       IF #enterAddress THEN

                           REGION "TURN OFF THE LIGHTS"
                               #enterAddress := FALSE;
                           END_REGION

                           REGION "ENTER PART REQUEST"
                               #stations.me[#i].partRequested[#j] := TRUE;
                           END_REGION

                           REGION "ADDRESS"
                               #requests.row[#pRow].address := #address;
                           END_REGION

                           REGION "LINE"
                               #requests.row[#pRow].tfLine.value := #stations.me[#i].line;
                           END_REGION

                           REGION "DROP ZONE"
                               #requests.row[#pRow].tfDropZone.value := USINT_TO_WSTRING(#stations.me[#i].dropZone);
                           END_REGION

                           REGION "PART NUMBER"
                               #requests.row[#pRow].tfPartNumber.value := #stations.me[#i].partNumbers[#j];
                           END_REGION

                           REGION "ELLAPSED TIME"
                               #requests.row[#pRow].tfTime.value := "Real to WString Timer"(#stations.me[#i].elapsedTime.partReq[#j]);
                           END_REGION

                           REGION "ROW POINTER"

                               REGION "INCREMENT"
                                   #pRow := #pRow + 1;
                               END_REGION

                               REGION "HIGH LIMIT ROLLOVER"
                                   IF #pRow > "partReqDataRowCount" THEN
                                       #pRow := 0;
                                   END_IF;
                               END_REGION

                           END_REGION

                       END_IF;
                   END_REGION

               END_FOR;
           END_REGION

       END_FOR;
   END_REGION
END_FUNCTION_BLOCK

FUNCTION_BLOCK "Remove Part Request"   // FB13, SCL
{ S7_Optimized_Access := 'TRUE' }
VERSION : 0.1
   VAR_IN_OUT
      pRow : Int;
      requests : "Part Request Data";
      stations : "Stations";
      reqCollapse : Bool;
   END_VAR
   VAR
      old : Struct
         partReq : "Station Old Presses";
      END_STRUCT;
   END_VAR
   VAR_TEMP
      address : UInt;
      blankRow : "Table Row";
      hasPart : Bool;
      i : Int;
      j : Int;
      k : Int;
      logAddress : UInt;
      noPart : Bool;
      oldPartReq : Bool;
      partNumber : WString;
      partReq : Bool;
      pRemoveRow : Int;
      removeAddress : Bool;
   END_VAR
BEGIN


   REGION "FOR EACH STATION"
       FOR #i := 0 TO "stnCount" DO

           REGION "FOR EACH BUTTON"
               FOR #j := 1 TO "ptsPerStn" DO

                   REGION "COPY TO LOCAL"
                       #partReq := #stations.me[#i].btnStates[#j];
                       #oldPartReq := #old.partReq.me[#i, #j];
                   END_REGION

                   REGION "DETERMINE STATE"

                       REGION "PART REQUEST FALLING EDGE"
                           IF NOT #partReq AND #oldPartReq THEN

                               REGION "COPY TO LOCAL"
                                   #partNumber := #stations.me[#i].partNumbers[#j];
                               END_REGION

                               REGION "BUTTON HAS NO PART"
                                   IF #partNumber = wstring#'' THEN
                                       #hasPart := FALSE;
                                       #noPart := TRUE;
                                   END_IF;
                               END_REGION

                               REGION "BUTTON HAS PART"
                                   IF #partNumber <> wstring#'' THEN
                                       #hasPart := TRUE;
                                       #noPart := FALSE;
                                   END_IF;
                               END_REGION

                           END_IF;

                           REGION "SAVE FOR CHANGE DETECTION"
                               #old.partReq.me[#i, #j] := #partReq;
                           END_REGION

                       END_REGION

                   END_REGION

                   REGION "NO PART"
                       IF #noPart THEN

                           REGION "TURN OFF THE LIGHTS"
                               #hasPart := FALSE;
                               #noPart := FALSE;
                           END_REGION

                       END_IF;

                   END_REGION

                   REGION "HAS PART"
                       IF #hasPart THEN

                           REGION "TURN OFF THE LIGHTS"
                               #hasPart := FALSE;
                           END_REGION

                           REGION "CALCULATE ADDRESS"
                               #address := (INT_TO_UINT(#i) + 1) * 10 + (INT_TO_UINT(#j) + 1);
                           END_REGION

                           REGION "RESET FLAG"
                               #removeAddress := FALSE;
                           END_REGION

                           REGION "SEARCH EACH ROW IN PART DB"
                               FOR #k := 0 TO "partReqDataRowCount" DO

                                   REGION "COPY TO LOCAL"
                                       #logAddress := #requests.row[#k].address;
                                   END_REGION

                                   REGION "ON MATCH"
                                       IF #logAddress = #address THEN

                                           REGION "SET FLAG"
                                               #removeAddress := TRUE;
                                           END_REGION

                                           REGION "SAVE POINTER"
                                               #pRemoveRow := #k;
                                           END_REGION

                                       END_IF;
                                   END_REGION

                               END_FOR;
                           END_REGION

                       END_IF;
                   END_REGION

                   REGION "REMOVE ADDRESS"
                       IF #removeAddress THEN

                           REGION "TURN OFF THE LIGHTS"
                               #removeAddress := FALSE;
                           END_REGION

                           REGION "TURN OFF REQUEST"
                               #stations.me[#i].partRequested[#j] := FALSE;
                           END_REGION

                           REGION "REMOVAL PROCESS"

                               REGION "REMOVE ROW"
                                   #requests.row[#pRemoveRow] := #blankRow;
                                   #reqCollapse := TRUE;
                               END_REGION

                               REGION "REMOVE PART ORDERED"
                                   #stations.me[#i].partOrdered[#j] := FALSE;
                               END_REGION

                           END_REGION

                           REGION "ROW POINTER"

